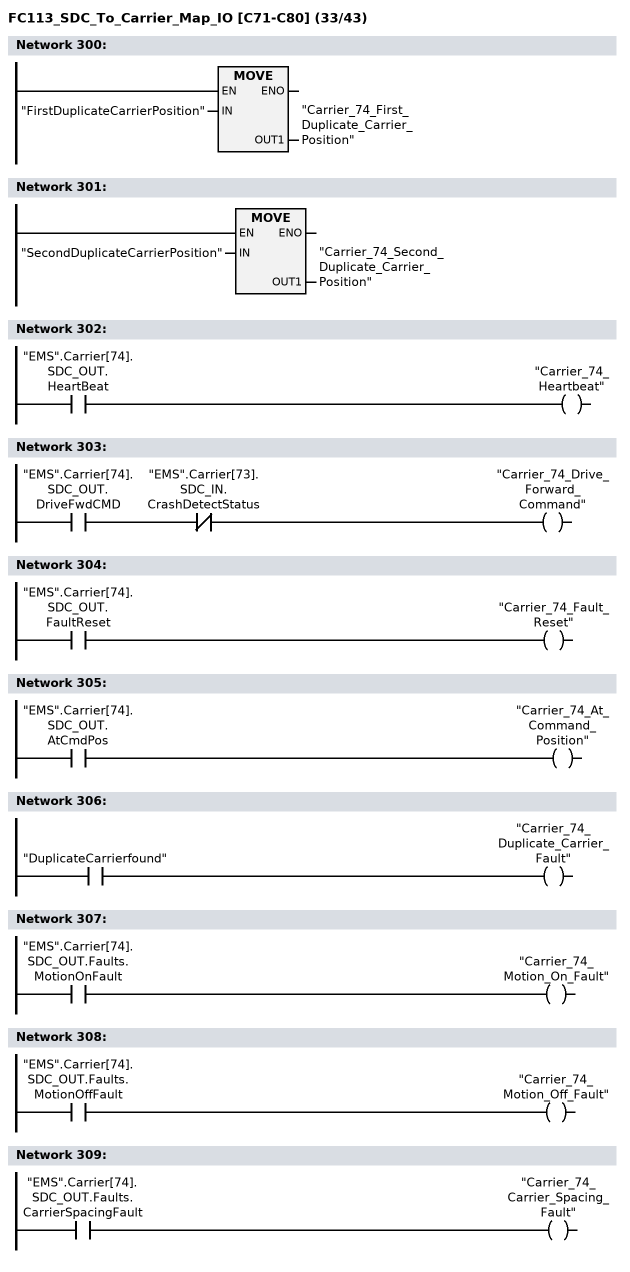
   RUNG wire#powerrail
      Move(in := "FirstDuplicateCarrierPosition", out1 => "Carrier_74_First_Duplicate_Carrier_Position")
   END_RUNG
   // the same network as SCL:
   "Carrier_74_First_Duplicate_Carrier_Position" := "FirstDuplicateCarrierPosition";
END_REGION

REGION Network 301
   RUNG wire#powerrail
      Move(in := "SecondDuplicateCarrierPosition", out1 => "Carrier_74_Second_Duplicate_Carrier_Position")
   END_RUNG
   // the same network as SCL:
   "Carrier_74_Second_Duplicate_Carrier_Position" := "SecondDuplicateCarrierPosition";
END_REGION

REGION Network 302
   RUNG wire#powerrail
      Contact( "EMS".Carrier[74].SDC_OUT.HeartBeat )
      Coil( "Carrier_74_Heartbeat" )
   END_RUNG
   // the same network as SCL:
   "Carrier_74_Heartbeat" := "EMS".Carrier[74].SDC_OUT.HeartBeat;
END_REGION

REGION Network 303
   RUNG wire#powerrail
      Contact( "EMS".Carrier[74].SDC_OUT.DriveFwdCMD )
      I_Contact( "EMS".Carrier[73].SDC_IN.CrashDetectStatus )
      Coil( "Carrier_74_Drive_Forward_Command" )
   END_RUNG
   // the same network as SCL:
   "Carrier_74_Drive_Forward_Command" := "EMS".Carrier[74].SDC_OUT.DriveFwdCMD AND NOT "EMS".Carrier[73].SDC_IN.CrashDetectStatus;
END_REGION

REGION Network 304
   RUNG wire#powerrail
      Contact( "EMS".Carrier[74].SDC_OUT.FaultReset )
      Coil( "Carrier_74_Fault_Reset" )
   END_RUNG
   // the same network as SCL:
   "Carrier_74_Fault_Reset" := "EMS".Carrier[74].SDC_OUT.FaultReset;
END_REGION

REGION Network 305
   RUNG wire#powerrail
      Contact( "EMS".Carrier[74].SDC_OUT.AtCmdPos )
      Coil( "Carrier_74_At_Command_Position" )
   END_RUNG
   // the same network as SCL:
   "Carrier_74_At_Command_Position" := "EMS".Carrier[74].SDC_OUT.AtCmdPos;
END_REGION

REGION Network 306
   RUNG wire#powerrail
      Contact( "DuplicateCarrierfound" )
      Coil( "Carrier_74_Duplicate_Carrier_Fault" )
   END_RUNG
   // the same network as SCL:
   "Carrier_74_Duplicate_Carrier_Fault" := "DuplicateCarrierfound";
END_REGION

REGION Network 307
   RUNG wire#powerrail
      Contact( "EMS".Carrier[74].SDC_OUT.Faults.MotionOnFault )
      Coil( "Carrier_74_Motion_On_Fault" )
   END_RUNG
   // the same network as SCL:
   "Carrier_74_Motion_On_Fault" := "EMS".Carrier[74].SDC_OUT.Faults.MotionOnFault;
END_REGION

REGION Network 308
   RUNG wire#powerrail
      Contact( "EMS".Carrier[74].SDC_OUT.Faults.MotionOffFault )
      Coil( "Carrier_74_Motion_Off_Fault" )
   END_RUNG
   // the same network as SCL:
   "Carrier_74_Motion_Off_Fault" := "EMS".Carrier[74].SDC_OUT.Faults.MotionOffFault;
END_REGION

REGION Network 309
   RUNG wire#powerrail
      Contact( "EMS".Carrier[74].SDC_OUT.Faults.CarrierSpacingFault )
      Coil( "Carrier_74_Carrier_Spacing_Fault" )
   END_RUNG
   // the same network as SCL:
   "Carrier_74_Carrier_Spacing_Fault" := "EMS".Carrier[74].SDC_OUT.Faults.CarrierSpacingFault;
END_REGION

REGION Network 310
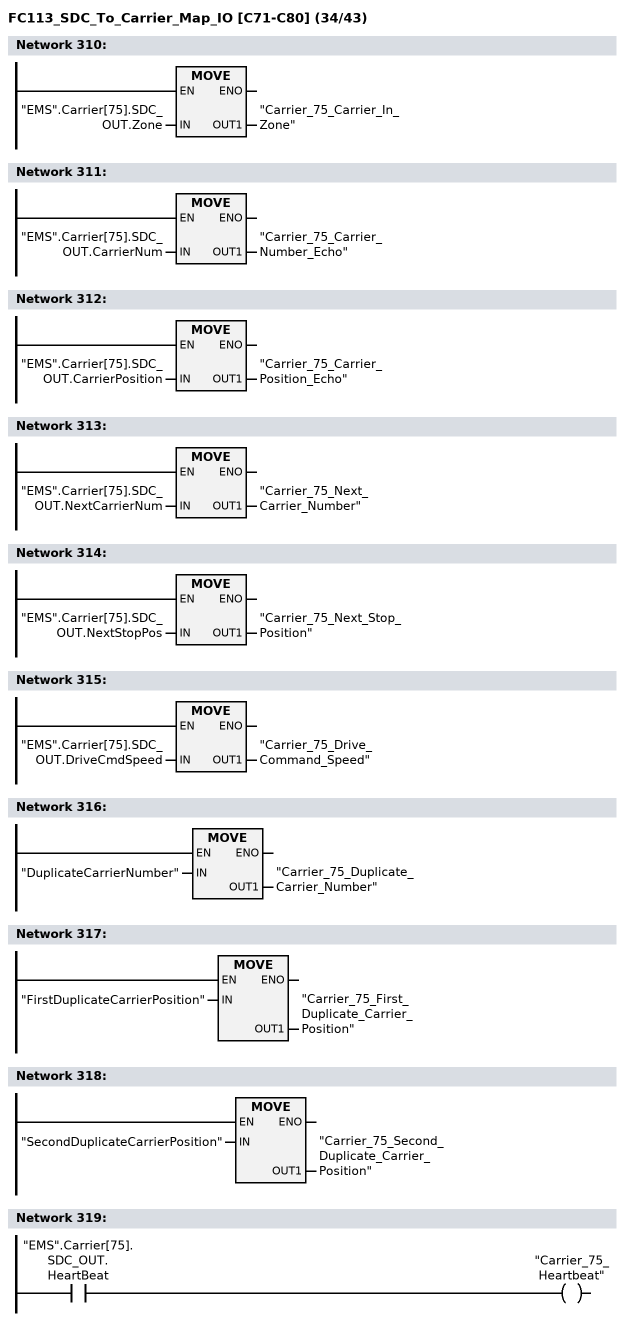
   RUNG wire#powerrail
      Move(in := "EMS".Carrier[75].SDC_OUT.Zone, out1 => "Carrier_75_Carrier_In_Zone")
   END_RUNG
   // the same network as SCL:
   "Carrier_75_Carrier_In_Zone" := "EMS".Carrier[75].SDC_OUT.Zone;
END_REGION

REGION Network 311
   RUNG wire#powerrail
      Move(in := "EMS".Carrier[75].SDC_OUT.CarrierNum, out1 => "Carrier_75_Carrier_Number_Echo")
   END_RUNG
   // the same network as SCL:
   "Carrier_75_Carrier_Number_Echo" := "EMS".Carrier[75].SDC_OUT.CarrierNum;
END_REGION

REGION Network 312
   RUNG wire#powerrail
      Move(in := "EMS".Carrier[75].SDC_OUT.CarrierPosition, out1 => "Carrier_75_Carrier_Position_Echo")
   END_RUNG
   // the same network as SCL:
   "Carrier_75_Carrier_Position_Echo" := "EMS".Carrier[75].SDC_OUT.CarrierPosition;
END_REGION

REGION Network 313
   RUNG wire#powerrail
      Move(in := "EMS".Carrier[75].SDC_OUT.NextCarrierNum, out1 => "Carrier_75_Next_Carrier_Number")
   END_RUNG
   // the same network as SCL:
   "Carrier_75_Next_Carrier_Number" := "EMS".Carrier[75].SDC_OUT.NextCarrierNum;
END_REGION

REGION Network 314
   RUNG wire#powerrail
      Move(in := "EMS".Carrier[75].SDC_OUT.NextStopPos, out1 => "Carrier_75_Next_Stop_Position")
   END_RUNG
   // the same network as SCL:
   "Carrier_75_Next_Stop_Position" := "EMS".Carrier[75].SDC_OUT.NextStopPos;
END_REGION

REGION Network 315
   RUNG wire#powerrail
      Move(in := "EMS".Carrier[75].SDC_OUT.DriveCmdSpeed, out1 => "Carrier_75_Drive_Command_Speed")
   END_RUNG
   // the same network as SCL:
   "Carrier_75_Drive_Command_Speed" := "EMS".Carrier[75].SDC_OUT.DriveCmdSpeed;
END_REGION

REGION Network 316
   RUNG wire#powerrail
      Move(in := "DuplicateCarrierNumber", out1 => "Carrier_75_Duplicate_Carrier_Number")
   END_RUNG
   // the same network as SCL:
   "Carrier_75_Duplicate_Carrier_Number" := "DuplicateCarrierNumber";
END_REGION

REGION Network 317
   RUNG wire#powerrail
      Move(in := "FirstDuplicateCarrierPosition", out1 => "Carrier_75_First_Duplicate_Carrier_Position")
   END_RUNG
   // the same network as SCL:
   "Carrier_75_First_Duplicate_Carrier_Position" := "FirstDuplicateCarrierPosition";
END_REGION

REGION Network 318
   RUNG wire#powerrail
      Move(in := "SecondDuplicateCarrierPosition", out1 => "Carrier_75_Second_Duplicate_Carrier_Position")
   END_RUNG
   // the same network as SCL:
   "Carrier_75_Second_Duplicate_Carrier_Position" := "SecondDuplicateCarrierPosition";
END_REGION

REGION Network 319
   RUNG wire#powerrail
      Contact( "EMS".Carrier[75].SDC_OUT.HeartBeat )
      Coil( "Carrier_75_Heartbeat" )
   END_RUNG
   // the same network as SCL:
   "Carrier_75_Heartbeat" := "EMS".Carrier[75].SDC_OUT.HeartBeat;
END_REGION

REGION Network 320
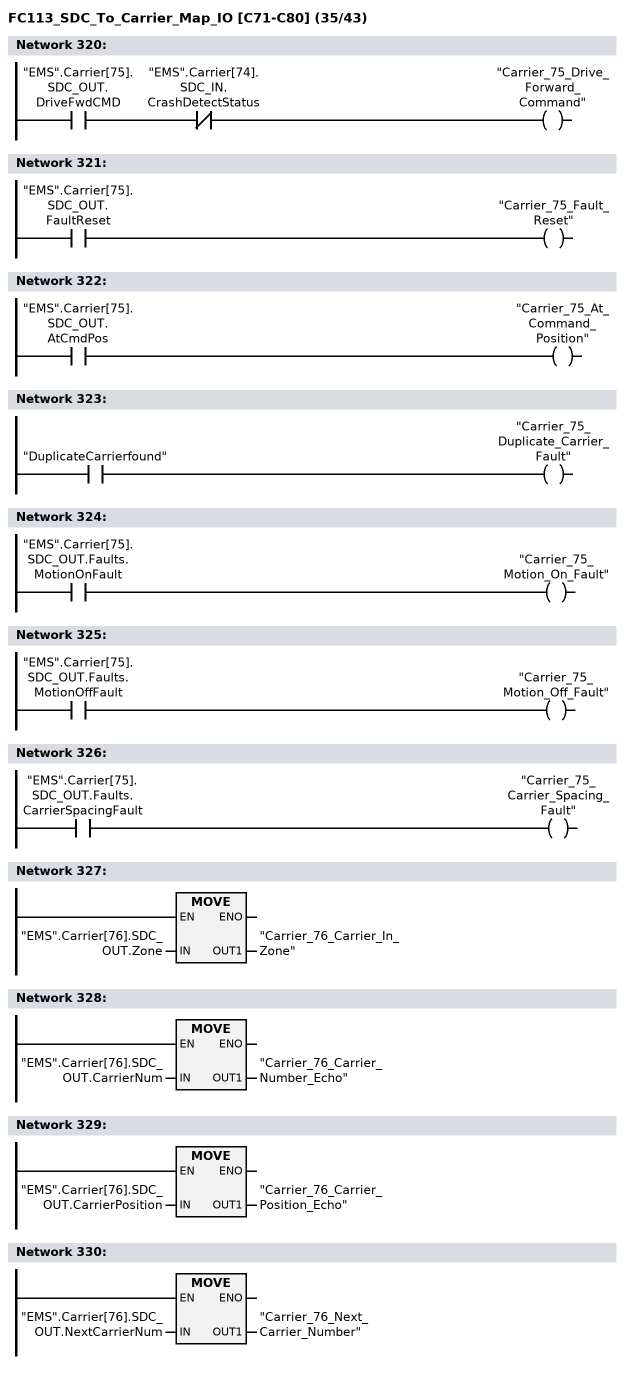
   RUNG wire#powerrail
      Contact( "EMS".Carrier[75].SDC_OUT.DriveFwdCMD )
      I_Contact( "EMS".Carrier[74].SDC_IN.CrashDetectStatus )
      Coil( "Carrier_75_Drive_Forward_Command" )
   END_RUNG
   // the same network as SCL:
   "Carrier_75_Drive_Forward_Command" := "EMS".Carrier[75].SDC_OUT.DriveFwdCMD AND NOT "EMS".Carrier[74].SDC_IN.CrashDetectStatus;
END_REGION

REGION Network 321
   RUNG wire#powerrail
      Contact( "EMS".Carrier[75].SDC_OUT.FaultReset )
      Coil( "Carrier_75_Fault_Reset" )
   END_RUNG
   // the same network as SCL:
   "Carrier_75_Fault_Reset" := "EMS".Carrier[75].SDC_OUT.FaultReset;
END_REGION

REGION Network 322
   RUNG wire#powerrail
      Contact( "EMS".Carrier[75].SDC_OUT.AtCmdPos )
      Coil( "Carrier_75_At_Command_Position" )
   END_RUNG
   // the same network as SCL:
   "Carrier_75_At_Command_Position" := "EMS".Carrier[75].SDC_OUT.AtCmdPos;
END_REGION

REGION Network 323
   RUNG wire#powerrail
      Contact( "DuplicateCarrierfound" )
      Coil( "Carrier_75_Duplicate_Carrier_Fault" )
   END_RUNG
   // the same network as SCL:
   "Carrier_75_Duplicate_Carrier_Fault" := "DuplicateCarrierfound";
END_REGION

REGION Network 324
   RUNG wire#powerrail
      Contact( "EMS".Carrier[75].SDC_OUT.Faults.MotionOnFault )
      Coil( "Carrier_75_Motion_On_Fault" )
   END_RUNG
   // the same network as SCL:
   "Carrier_75_Motion_On_Fault" := "EMS".Carrier[75].SDC_OUT.Faults.MotionOnFault;
END_REGION

REGION Network 325
   RUNG wire#powerrail
      Contact( "EMS".Carrier[75].SDC_OUT.Faults.MotionOffFault )
      Coil( "Carrier_75_Motion_Off_Fault" )
   END_RUNG
   // the same network as SCL:
   "Carrier_75_Motion_Off_Fault" := "EMS".Carrier[75].SDC_OUT.Faults.MotionOffFault;
END_REGION

REGION Network 326
   RUNG wire#powerrail
      Contact( "EMS".Carrier[75].SDC_OUT.Faults.CarrierSpacingFault )
      Coil( "Carrier_75_Carrier_Spacing_Fault" )
   END_RUNG
   // the same network as SCL:
   "Carrier_75_Carrier_Spacing_Fault" := "EMS".Carrier[75].SDC_OUT.Faults.CarrierSpacingFault;
END_REGION

REGION Network 327
   RUNG wire#powerrail
      Move(in := "EMS".Carrier[76].SDC_OUT.Zone, out1 => "Carrier_76_Carrier_In_Zone")
   END_RUNG
   // the same network as SCL:
   "Carrier_76_Carrier_In_Zone" := "EMS".Carrier[76].SDC_OUT.Zone;
END_REGION

REGION Network 328
   RUNG wire#powerrail
      Move(in := "EMS".Carrier[76].SDC_OUT.CarrierNum, out1 => "Carrier_76_Carrier_Number_Echo")
   END_RUNG
   // the same network as SCL:
   "Carrier_76_Carrier_Number_Echo" := "EMS".Carrier[76].SDC_OUT.CarrierNum;
END_REGION

REGION Network 329
   RUNG wire#powerrail
      Move(in := "EMS".Carrier[76].SDC_OUT.CarrierPosition, out1 => "Carrier_76_Carrier_Position_Echo")
   END_RUNG
   // the same network as SCL:
   "Carrier_76_Carrier_Position_Echo" := "EMS".Carrier[76].SDC_OUT.CarrierPosition;
END_REGION

REGION Network 330
   RUNG wire#powerrail
      Move(in := "EMS".Carrier[76].SDC_OUT.NextCarrierNum, out1 => "Carrier_76_Next_Carrier_Number")
   END_RUNG
   // the same network as SCL:
   "Carrier_76_Next_Carrier_Number" := "EMS".Carrier[76].SDC_OUT.NextCarrierNum;
END_REGION

REGION Network 331
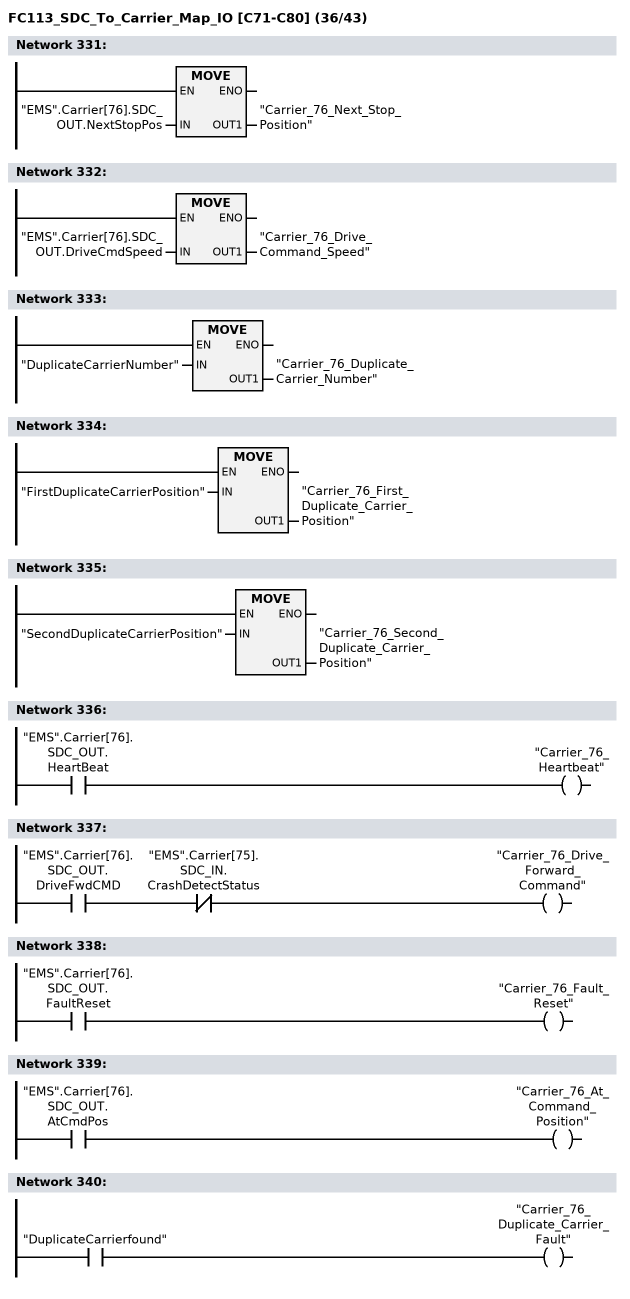
   RUNG wire#powerrail
      Move(in := "EMS".Carrier[76].SDC_OUT.NextStopPos, out1 => "Carrier_76_Next_Stop_Position")
   END_RUNG
   // the same network as SCL:
   "Carrier_76_Next_Stop_Position" := "EMS".Carrier[76].SDC_OUT.NextStopPos;
END_REGION

REGION Network 332
   RUNG wire#powerrail
      Move(in := "EMS".Carrier[76].SDC_OUT.DriveCmdSpeed, out1 => "Carrier_76_Drive_Command_Speed")
   END_RUNG
   // the same network as SCL:
   "Carrier_76_Drive_Command_Speed" := "EMS".Carrier[76].SDC_OUT.DriveCmdSpeed;
END_REGION

REGION Network 333
   RUNG wire#powerrail
      Move(in := "DuplicateCarrierNumber", out1 => "Carrier_76_Duplicate_Carrier_Number")
   END_RUNG
   // the same network as SCL:
   "Carrier_76_Duplicate_Carrier_Number" := "DuplicateCarrierNumber";
END_REGION

REGION Network 334
   RUNG wire#powerrail
      Move(in := "FirstDuplicateCarrierPosition", out1 => "Carrier_76_First_Duplicate_Carrier_Position")
   END_RUNG
   // the same network as SCL:
   "Carrier_76_First_Duplicate_Carrier_Position" := "FirstDuplicateCarrierPosition";
END_REGION

REGION Network 335
   RUNG wire#powerrail
      Move(in := "SecondDuplicateCarrierPosition", out1 => "Carrier_76_Second_Duplicate_Carrier_Position")
   END_RUNG
   // the same network as SCL:
   "Carrier_76_Second_Duplicate_Carrier_Position" := "SecondDuplicateCarrierPosition";
END_REGION

REGION Network 336
   RUNG wire#powerrail
      Contact( "EMS".Carrier[76].SDC_OUT.HeartBeat )
      Coil( "Carrier_76_Heartbeat" )
   END_RUNG
   // the same network as SCL:
   "Carrier_76_Heartbeat" := "EMS".Carrier[76].SDC_OUT.HeartBeat;
END_REGION

REGION Network 337
   RUNG wire#powerrail
      Contact( "EMS".Carrier[76].SDC_OUT.DriveFwdCMD )
      I_Contact( "EMS".Carrier[75].SDC_IN.CrashDetectStatus )
      Coil( "Carrier_76_Drive_Forward_Command" )
   END_RUNG
   // the same network as SCL:
   "Carrier_76_Drive_Forward_Command" := "EMS".Carrier[76].SDC_OUT.DriveFwdCMD AND NOT "EMS".Carrier[75].SDC_IN.CrashDetectStatus;
END_REGION

REGION Network 338
   RUNG wire#powerrail
      Contact( "EMS".Carrier[76].SDC_OUT.FaultReset )
      Coil( "Carrier_76_Fault_Reset" )
   END_RUNG
   // the same network as SCL:
   "Carrier_76_Fault_Reset" := "EMS".Carrier[76].SDC_OUT.FaultReset;
END_REGION

REGION Network 339
   RUNG wire#powerrail
      Contact( "EMS".Carrier[76].SDC_OUT.AtCmdPos )
      Coil( "Carrier_76_At_Command_Position" )
   END_RUNG
   // the same network as SCL:
   "Carrier_76_At_Command_Position" := "EMS".Carrier[76].SDC_OUT.AtCmdPos;
END_REGION

REGION Network 340
   RUNG wire#powerrail
      Contact( "DuplicateCarrierfound" )
      Coil( "Carrier_76_Duplicate_Carrier_Fault" )
   END_RUNG
   // the same network as SCL:
   "Carrier_76_Duplicate_Carrier_Fault" := "DuplicateCarrierfound";
END_REGION

REGION Network 341
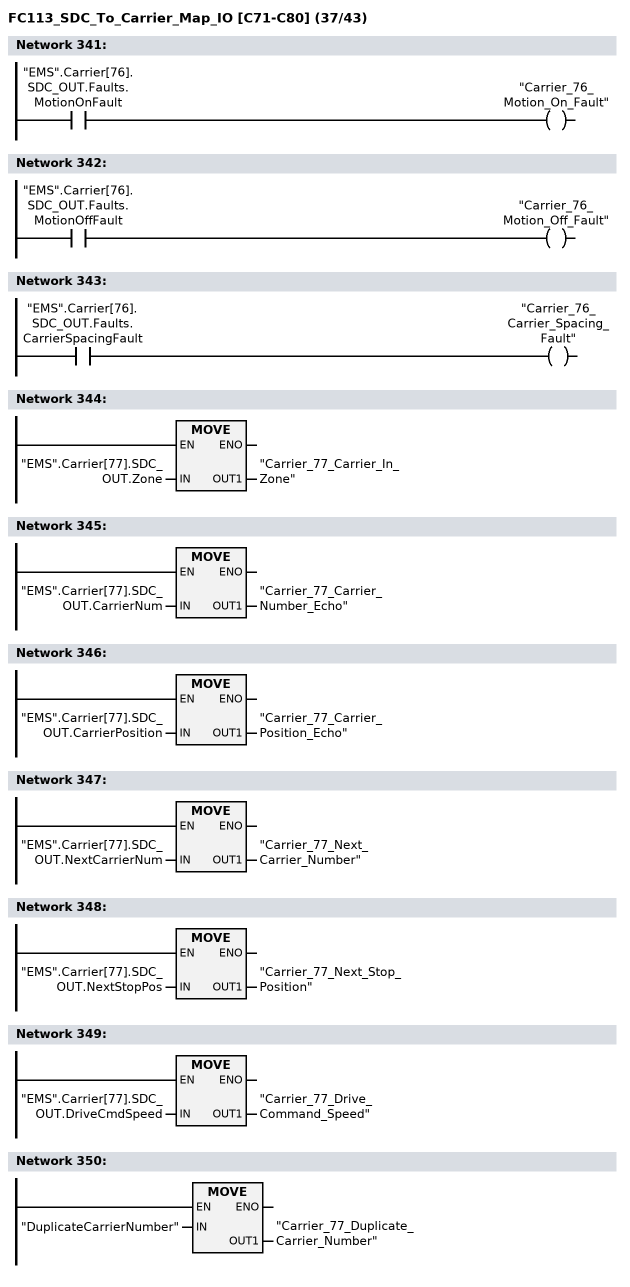
   RUNG wire#powerrail
      Contact( "EMS".Carrier[76].SDC_OUT.Faults.MotionOnFault )
      Coil( "Carrier_76_Motion_On_Fault" )
   END_RUNG
   // the same network as SCL:
   "Carrier_76_Motion_On_Fault" := "EMS".Carrier[76].SDC_OUT.Faults.MotionOnFault;
END_REGION

REGION Network 342
   RUNG wire#powerrail
      Contact( "EMS".Carrier[76].SDC_OUT.Faults.MotionOffFault )
      Coil( "Carrier_76_Motion_Off_Fault" )
   END_RUNG
   // the same network as SCL:
   "Carrier_76_Motion_Off_Fault" := "EMS".Carrier[76].SDC_OUT.Faults.MotionOffFault;
END_REGION

REGION Network 343
   RUNG wire#powerrail
      Contact( "EMS".Carrier[76].SDC_OUT.Faults.CarrierSpacingFault )
      Coil( "Carrier_76_Carrier_Spacing_Fault" )
   END_RUNG
   // the same network as SCL:
   "Carrier_76_Carrier_Spacing_Fault" := "EMS".Carrier[76].SDC_OUT.Faults.CarrierSpacingFault;
END_REGION

REGION Network 344
   RUNG wire#powerrail
      Move(in := "EMS".Carrier[77].SDC_OUT.Zone, out1 => "Carrier_77_Carrier_In_Zone")
   END_RUNG
   // the same network as SCL:
   "Carrier_77_Carrier_In_Zone" := "EMS".Carrier[77].SDC_OUT.Zone;
END_REGION

REGION Network 345
   RUNG wire#powerrail
      Move(in := "EMS".Carrier[77].SDC_OUT.CarrierNum, out1 => "Carrier_77_Carrier_Number_Echo")
   END_RUNG
   // the same network as SCL:
   "Carrier_77_Carrier_Number_Echo" := "EMS".Carrier[77].SDC_OUT.CarrierNum;
END_REGION

REGION Network 346
   RUNG wire#powerrail
      Move(in := "EMS".Carrier[77].SDC_OUT.CarrierPosition, out1 => "Carrier_77_Carrier_Position_Echo")
   END_RUNG
   // the same network as SCL:
   "Carrier_77_Carrier_Position_Echo" := "EMS".Carrier[77].SDC_OUT.CarrierPosition;
END_REGION

REGION Network 347
   RUNG wire#powerrail
      Move(in := "EMS".Carrier[77].SDC_OUT.NextCarrierNum, out1 => "Carrier_77_Next_Carrier_Number")
   END_RUNG
   // the same network as SCL:
   "Carrier_77_Next_Carrier_Number" := "EMS".Carrier[77].SDC_OUT.NextCarrierNum;
END_REGION

REGION Network 348
   RUNG wire#powerrail
      Move(in := "EMS".Carrier[77].SDC_OUT.NextStopPos, out1 => "Carrier_77_Next_Stop_Position")
   END_RUNG
   // the same network as SCL:
   "Carrier_77_Next_Stop_Position" := "EMS".Carrier[77].SDC_OUT.NextStopPos;
END_REGION

REGION Network 349
   RUNG wire#powerrail
      Move(in := "EMS".Carrier[77].SDC_OUT.DriveCmdSpeed, out1 => "Carrier_77_Drive_Command_Speed")
   END_RUNG
   // the same network as SCL:
   "Carrier_77_Drive_Command_Speed" := "EMS".Carrier[77].SDC_OUT.DriveCmdSpeed;
END_REGION

REGION Network 350
   RUNG wire#powerrail
      Move(in := "DuplicateCarrierNumber", out1 => "Carrier_77_Duplicate_Carrier_Number")
   END_RUNG
   // the same network as SCL:
   "Carrier_77_Duplicate_Carrier_Number" := "DuplicateCarrierNumber";
END_REGION

REGION Network 351
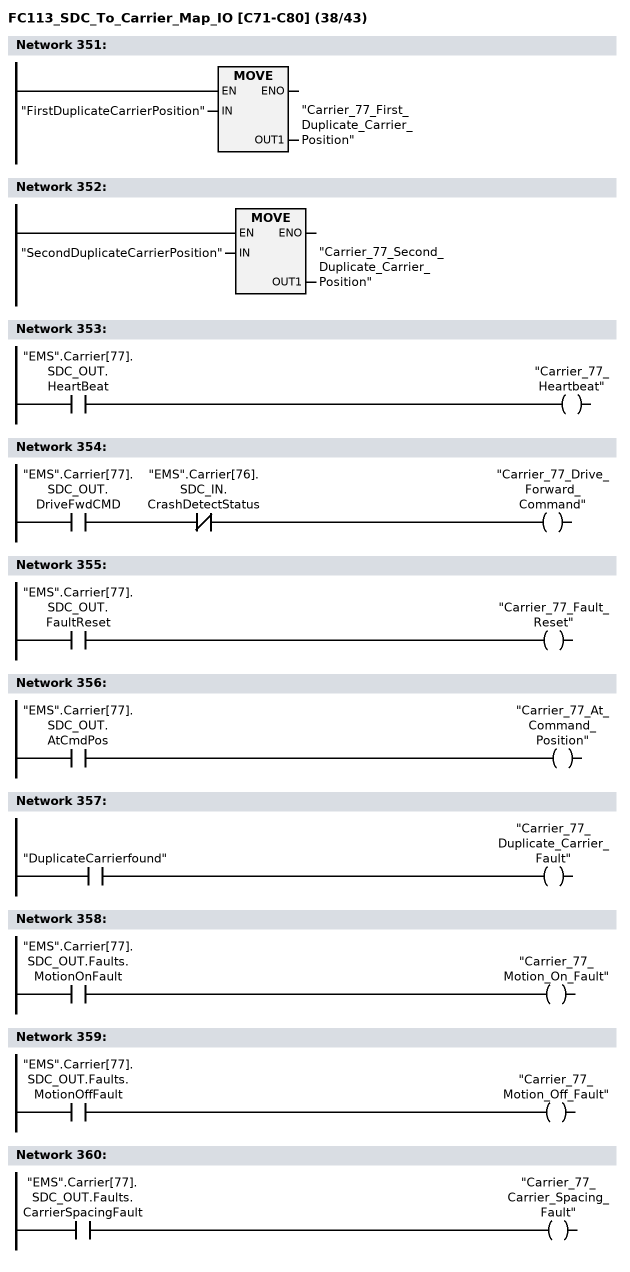
   RUNG wire#powerrail
      Move(in := "FirstDuplicateCarrierPosition", out1 => "Carrier_77_First_Duplicate_Carrier_Position")
   END_RUNG
   // the same network as SCL:
   "Carrier_77_First_Duplicate_Carrier_Position" := "FirstDuplicateCarrierPosition";
END_REGION

REGION Network 352
   RUNG wire#powerrail
      Move(in := "SecondDuplicateCarrierPosition", out1 => "Carrier_77_Second_Duplicate_Carrier_Position")
   END_RUNG
   // the same network as SCL:
   "Carrier_77_Second_Duplicate_Carrier_Position" := "SecondDuplicateCarrierPosition";
END_REGION

REGION Network 353
   RUNG wire#powerrail
      Contact( "EMS".Carrier[77].SDC_OUT.HeartBeat )
      Coil( "Carrier_77_Heartbeat" )
   END_RUNG
   // the same network as SCL:
   "Carrier_77_Heartbeat" := "EMS".Carrier[77].SDC_OUT.HeartBeat;
END_REGION

REGION Network 354
   RUNG wire#powerrail
      Contact( "EMS".Carrier[77].SDC_OUT.DriveFwdCMD )
      I_Contact( "EMS".Carrier[76].SDC_IN.CrashDetectStatus )
      Coil( "Carrier_77_Drive_Forward_Command" )
   END_RUNG
   // the same network as SCL:
   "Carrier_77_Drive_Forward_Command" := "EMS".Carrier[77].SDC_OUT.DriveFwdCMD AND NOT "EMS".Carrier[76].SDC_IN.CrashDetectStatus;
END_REGION

REGION Network 355
   RUNG wire#powerrail
      Contact( "EMS".Carrier[77].SDC_OUT.FaultReset )
      Coil( "Carrier_77_Fault_Reset" )
   END_RUNG
   // the same network as SCL:
   "Carrier_77_Fault_Reset" := "EMS".Carrier[77].SDC_OUT.FaultReset;
END_REGION

REGION Network 356
   RUNG wire#powerrail
      Contact( "EMS".Carrier[77].SDC_OUT.AtCmdPos )
      Coil( "Carrier_77_At_Command_Position" )
   END_RUNG
   // the same network as SCL:
   "Carrier_77_At_Command_Position" := "EMS".Carrier[77].SDC_OUT.AtCmdPos;
END_REGION

REGION Network 357
   RUNG wire#powerrail
      Contact( "DuplicateCarrierfound" )
      Coil( "Carrier_77_Duplicate_Carrier_Fault" )
   END_RUNG
   // the same network as SCL:
   "Carrier_77_Duplicate_Carrier_Fault" := "DuplicateCarrierfound";
END_REGION

REGION Network 358
   RUNG wire#powerrail
      Contact( "EMS".Carrier[77].SDC_OUT.Faults.MotionOnFault )
      Coil( "Carrier_77_Motion_On_Fault" )
   END_RUNG
   // the same network as SCL:
   "Carrier_77_Motion_On_Fault" := "EMS".Carrier[77].SDC_OUT.Faults.MotionOnFault;
END_REGION

REGION Network 359
   RUNG wire#powerrail
      Contact( "EMS".Carrier[77].SDC_OUT.Faults.MotionOffFault )
      Coil( "Carrier_77_Motion_Off_Fault" )
   END_RUNG
   // the same network as SCL:
   "Carrier_77_Motion_Off_Fault" := "EMS".Carrier[77].SDC_OUT.Faults.MotionOffFault;
END_REGION

REGION Network 360
   RUNG wire#powerrail
      Contact( "EMS".Carrier[77].SDC_OUT.Faults.CarrierSpacingFault )
      Coil( "Carrier_77_Carrier_Spacing_Fault" )
   END_RUNG
   // the same network as SCL:
   "Carrier_77_Carrier_Spacing_Fault" := "EMS".Carrier[77].SDC_OUT.Faults.CarrierSpacingFault;
END_REGION

REGION Network 361
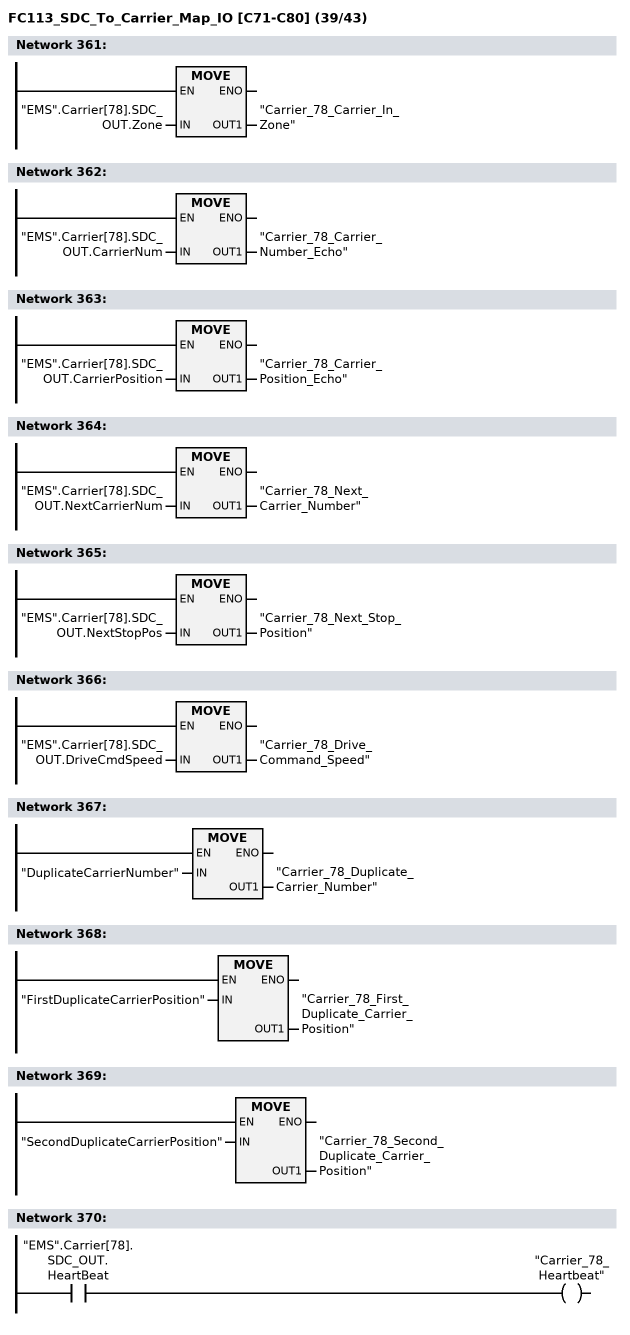
   RUNG wire#powerrail
      Move(in := "EMS".Carrier[78].SDC_OUT.Zone, out1 => "Carrier_78_Carrier_In_Zone")
   END_RUNG
   // the same network as SCL:
   "Carrier_78_Carrier_In_Zone" := "EMS".Carrier[78].SDC_OUT.Zone;
END_REGION

REGION Network 362
   RUNG wire#powerrail
      Move(in := "EMS".Carrier[78].SDC_OUT.CarrierNum, out1 => "Carrier_78_Carrier_Number_Echo")
   END_RUNG
   // the same network as SCL:
   "Carrier_78_Carrier_Number_Echo" := "EMS".Carrier[78].SDC_OUT.CarrierNum;
END_REGION

REGION Network 363
   RUNG wire#powerrail
      Move(in := "EMS".Carrier[78].SDC_OUT.CarrierPosition, out1 => "Carrier_78_Carrier_Position_Echo")
   END_RUNG
   // the same network as SCL:
   "Carrier_78_Carrier_Position_Echo" := "EMS".Carrier[78].SDC_OUT.CarrierPosition;
END_REGION

REGION Network 364
   RUNG wire#powerrail
      Move(in := "EMS".Carrier[78].SDC_OUT.NextCarrierNum, out1 => "Carrier_78_Next_Carrier_Number")
   END_RUNG
   // the same network as SCL:
   "Carrier_78_Next_Carrier_Number" := "EMS".Carrier[78].SDC_OUT.NextCarrierNum;
END_REGION

REGION Network 365
   RUNG wire#powerrail
      Move(in := "EMS".Carrier[78].SDC_OUT.NextStopPos, out1 => "Carrier_78_Next_Stop_Position")
   END_RUNG
   // the same network as SCL:
   "Carrier_78_Next_Stop_Position" := "EMS".Carrier[78].SDC_OUT.NextStopPos;
END_REGION

REGION Network 366
   RUNG wire#powerrail
      Move(in := "EMS".Carrier[78].SDC_OUT.DriveCmdSpeed, out1 => "Carrier_78_Drive_Command_Speed")
   END_RUNG
   // the same network as SCL:
   "Carrier_78_Drive_Command_Speed" := "EMS".Carrier[78].SDC_OUT.DriveCmdSpeed;
END_REGION

REGION Network 367
   RUNG wire#powerrail
      Move(in := "DuplicateCarrierNumber", out1 => "Carrier_78_Duplicate_Carrier_Number")
   END_RUNG
   // the same network as SCL:
   "Carrier_78_Duplicate_Carrier_Number" := "DuplicateCarrierNumber";
END_REGION

REGION Network 368
   RUNG wire#powerrail
      Move(in := "FirstDuplicateCarrierPosition", out1 => "Carrier_78_First_Duplicate_Carrier_Position")
   END_RUNG
   // the same network as SCL:
   "Carrier_78_First_Duplicate_Carrier_Position" := "FirstDuplicateCarrierPosition";
END_REGION

REGION Network 369
   RUNG wire#powerrail
      Move(in := "SecondDuplicateCarrierPosition", out1 => "Carrier_78_Second_Duplicate_Carrier_Position")
   END_RUNG
   // the same network as SCL:
   "Carrier_78_Second_Duplicate_Carrier_Position" := "SecondDuplicateCarrierPosition";
END_REGION

REGION Network 370
   RUNG wire#powerrail
      Contact( "EMS".Carrier[78].SDC_OUT.HeartBeat )
      Coil( "Carrier_78_Heartbeat" )
   END_RUNG
   // the same network as SCL:
   "Carrier_78_Heartbeat" := "EMS".Carrier[78].SDC_OUT.HeartBeat;
END_REGION

REGION Network 371
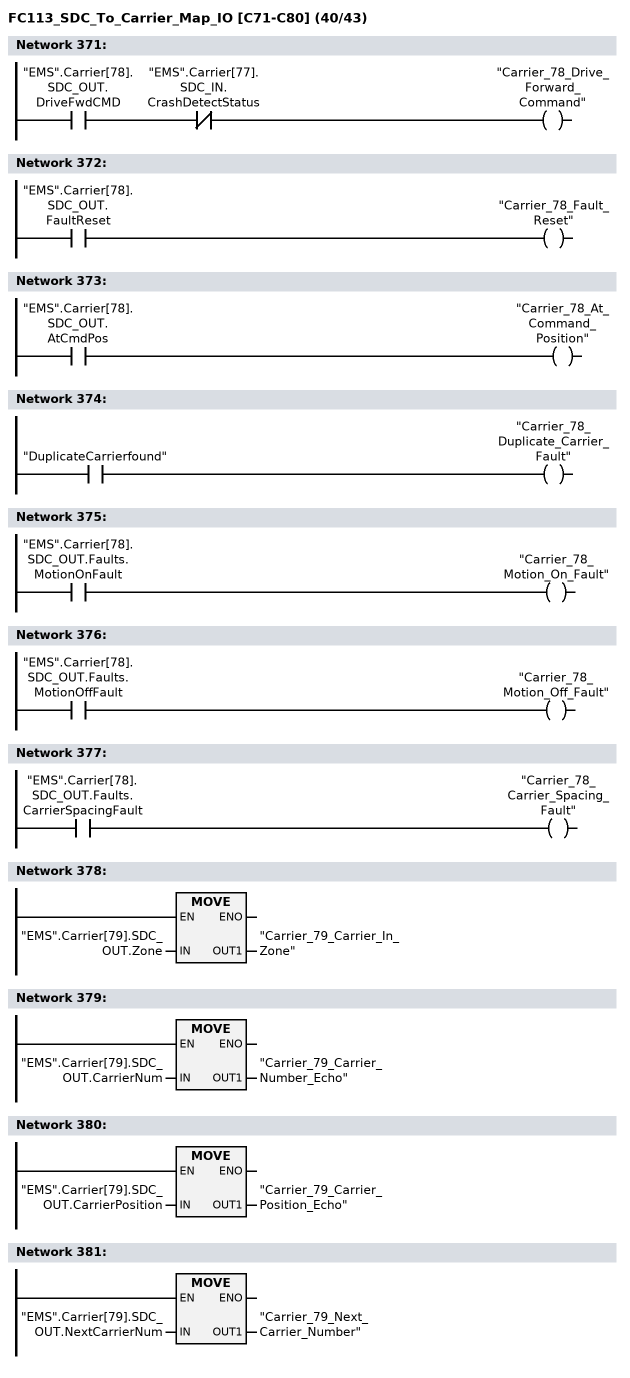
   RUNG wire#powerrail
      Contact( "EMS".Carrier[78].SDC_OUT.DriveFwdCMD )
      I_Contact( "EMS".Carrier[77].SDC_IN.CrashDetectStatus )
      Coil( "Carrier_78_Drive_Forward_Command" )
   END_RUNG
   // the same network as SCL:
   "Carrier_78_Drive_Forward_Command" := "EMS".Carrier[78].SDC_OUT.DriveFwdCMD AND NOT "EMS".Carrier[77].SDC_IN.CrashDetectStatus;
END_REGION

REGION Network 372
   RUNG wire#powerrail
      Contact( "EMS".Carrier[78].SDC_OUT.FaultReset )
      Coil( "Carrier_78_Fault_Reset" )
   END_RUNG
   // the same network as SCL:
   "Carrier_78_Fault_Reset" := "EMS".Carrier[78].SDC_OUT.FaultReset;
END_REGION

REGION Network 373
   RUNG wire#powerrail
      Contact( "EMS".Carrier[78].SDC_OUT.AtCmdPos )
      Coil( "Carrier_78_At_Command_Position" )
   END_RUNG
   // the same network as SCL:
   "Carrier_78_At_Command_Position" := "EMS".Carrier[78].SDC_OUT.AtCmdPos;
END_REGION

REGION Network 374
   RUNG wire#powerrail
      Contact( "DuplicateCarrierfound" )
      Coil( "Carrier_78_Duplicate_Carrier_Fault" )
   END_RUNG
   // the same network as SCL:
   "Carrier_78_Duplicate_Carrier_Fault" := "DuplicateCarrierfound";
END_REGION

REGION Network 375
   RUNG wire#powerrail
      Contact( "EMS".Carrier[78].SDC_OUT.Faults.MotionOnFault )
      Coil( "Carrier_78_Motion_On_Fault" )
   END_RUNG
   // the same network as SCL:
   "Carrier_78_Motion_On_Fault" := "EMS".Carrier[78].SDC_OUT.Faults.MotionOnFault;
END_REGION

REGION Network 376
   RUNG wire#powerrail
      Contact( "EMS".Carrier[78].SDC_OUT.Faults.MotionOffFault )
      Coil( "Carrier_78_Motion_Off_Fault" )
   END_RUNG
   // the same network as SCL:
   "Carrier_78_Motion_Off_Fault" := "EMS".Carrier[78].SDC_OUT.Faults.MotionOffFault;
END_REGION

REGION Network 377
   RUNG wire#powerrail
      Contact( "EMS".Carrier[78].SDC_OUT.Faults.CarrierSpacingFault )
      Coil( "Carrier_78_Carrier_Spacing_Fault" )
   END_RUNG
   // the same network as SCL:
   "Carrier_78_Carrier_Spacing_Fault" := "EMS".Carrier[78].SDC_OUT.Faults.CarrierSpacingFault;
END_REGION

REGION Network 378
   RUNG wire#powerrail
      Move(in := "EMS".Carrier[79].SDC_OUT.Zone, out1 => "Carrier_79_Carrier_In_Zone")
   END_RUNG
   // the same network as SCL:
   "Carrier_79_Carrier_In_Zone" := "EMS".Carrier[79].SDC_OUT.Zone;
END_REGION

REGION Network 379
   RUNG wire#powerrail
      Move(in := "EMS".Carrier[79].SDC_OUT.CarrierNum, out1 => "Carrier_79_Carrier_Number_Echo")
   END_RUNG
   // the same network as SCL:
   "Carrier_79_Carrier_Number_Echo" := "EMS".Carrier[79].SDC_OUT.CarrierNum;
END_REGION

REGION Network 380
   RUNG wire#powerrail
      Move(in := "EMS".Carrier[79].SDC_OUT.CarrierPosition, out1 => "Carrier_79_Carrier_Position_Echo")
   END_RUNG
   // the same network as SCL:
   "Carrier_79_Carrier_Position_Echo" := "EMS".Carrier[79].SDC_OUT.CarrierPosition;
END_REGION

REGION Network 381
   RUNG wire#powerrail
      Move(in := "EMS".Carrier[79].SDC_OUT.NextCarrierNum, out1 => "Carrier_79_Next_Carrier_Number")
   END_RUNG
   // the same network as SCL:
   "Carrier_79_Next_Carrier_Number" := "EMS".Carrier[79].SDC_OUT.NextCarrierNum;
END_REGION

REGION Network 382
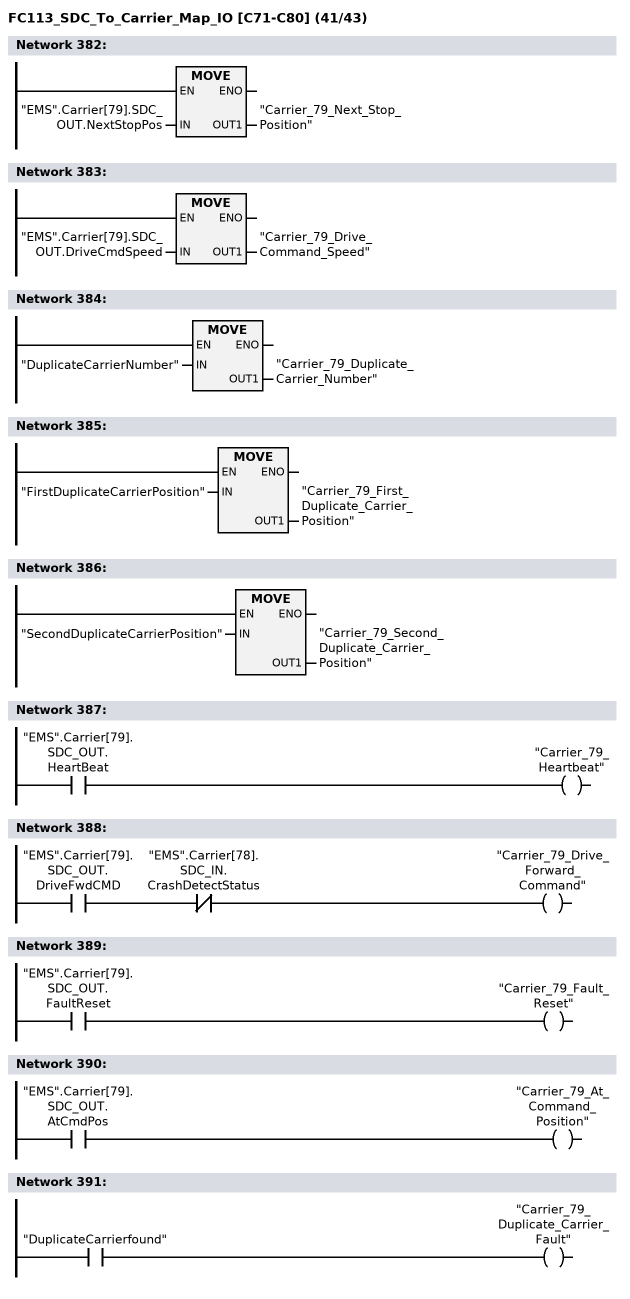
   RUNG wire#powerrail
      Move(in := "EMS".Carrier[79].SDC_OUT.NextStopPos, out1 => "Carrier_79_Next_Stop_Position")
   END_RUNG
   // the same network as SCL:
   "Carrier_79_Next_Stop_Position" := "EMS".Carrier[79].SDC_OUT.NextStopPos;
END_REGION

REGION Network 383
   RUNG wire#powerrail
      Move(in := "EMS".Carrier[79].SDC_OUT.DriveCmdSpeed, out1 => "Carrier_79_Drive_Command_Speed")
   END_RUNG
   // the same network as SCL:
   "Carrier_79_Drive_Command_Speed" := "EMS".Carrier[79].SDC_OUT.DriveCmdSpeed;
END_REGION

REGION Network 384
   RUNG wire#powerrail
      Move(in := "DuplicateCarrierNumber", out1 => "Carrier_79_Duplicate_Carrier_Number")
   END_RUNG
   // the same network as SCL:
   "Carrier_79_Duplicate_Carrier_Number" := "DuplicateCarrierNumber";
END_REGION

REGION Network 385
   RUNG wire#powerrail
      Move(in := "FirstDuplicateCarrierPosition", out1 => "Carrier_79_First_Duplicate_Carrier_Position")
   END_RUNG
   // the same network as SCL:
   "Carrier_79_First_Duplicate_Carrier_Position" := "FirstDuplicateCarrierPosition";
END_REGION

REGION Network 386
   RUNG wire#powerrail
      Move(in := "SecondDuplicateCarrierPosition", out1 => "Carrier_79_Second_Duplicate_Carrier_Position")
   END_RUNG
   // the same network as SCL:
   "Carrier_79_Second_Duplicate_Carrier_Position" := "SecondDuplicateCarrierPosition";
END_REGION

REGION Network 387
   RUNG wire#powerrail
      Contact( "EMS".Carrier[79].SDC_OUT.HeartBeat )
      Coil( "Carrier_79_Heartbeat" )
   END_RUNG
   // the same network as SCL:
   "Carrier_79_Heartbeat" := "EMS".Carrier[79].SDC_OUT.HeartBeat;
END_REGION

REGION Network 388
   RUNG wire#powerrail
      Contact( "EMS".Carrier[79].SDC_OUT.DriveFwdCMD )
      I_Contact( "EMS".Carrier[78].SDC_IN.CrashDetectStatus )
      Coil( "Carrier_79_Drive_Forward_Command" )
   END_RUNG
   // the same network as SCL:
   "Carrier_79_Drive_Forward_Command" := "EMS".Carrier[79].SDC_OUT.DriveFwdCMD AND NOT "EMS".Carrier[78].SDC_IN.CrashDetectStatus;
END_REGION

REGION Network 389
   RUNG wire#powerrail
      Contact( "EMS".Carrier[79].SDC_OUT.FaultReset )
      Coil( "Carrier_79_Fault_Reset" )
   END_RUNG
   // the same network as SCL:
   "Carrier_79_Fault_Reset" := "EMS".Carrier[79].SDC_OUT.FaultReset;
END_REGION

REGION Network 390
   RUNG wire#powerrail
      Contact( "EMS".Carrier[79].SDC_OUT.AtCmdPos )
      Coil( "Carrier_79_At_Command_Position" )
   END_RUNG
   // the same network as SCL:
   "Carrier_79_At_Command_Position" := "EMS".Carrier[79].SDC_OUT.AtCmdPos;
END_REGION

REGION Network 391
   RUNG wire#powerrail
      Contact( "DuplicateCarrierfound" )
      Coil( "Carrier_79_Duplicate_Carrier_Fault" )
   END_RUNG
   // the same network as SCL:
   "Carrier_79_Duplicate_Carrier_Fault" := "DuplicateCarrierfound";
END_REGION

REGION Network 392